HMI tags "Do_PLC"
   "System_okien_auto" : Bool = PLC HMI.System_okien_auto, 500 ms
   "Stopien_zasloniecia_rolet_manual" : Int = PLC HMI.Stopien_zasloniecia_rolet_manual, 100 ms
   "Przycisk_zraszania_manual" : Bool = PLC HMI.Przycisk_zraszacze_manual AT %Q0.2, 100 ms
   "Przycisk_wentylacja_manual" : Bool = PLC HMI.Przycisk_wentylacja_manual AT %Q0.1, 100 ms
   "Przycisk_grzanie_manual" : Bool = PLC HMI.Przycisk_grzanie_manual AT %Q0.0, 100 ms
   "Otwarcie_okien_man" : Bool = PLC HMI.Otwarcie_okien_manual AT %DB1.DBW0, 100 ms
   "Temperatura_auto" : Real = PLC HMI.Temperatura_auto, 500 ms
   "Naslonecznienie_auto" : Int = PLC HMI.Naslonecznienie_auto AT %DB1.DBW0, 500 ms
   "Wilgotnosc_powietrza_auto" : Int = PLC HMI.Wilgotnosc_powietrza_auto AT %DB1.DBW0, 500 ms
   "Wilgotnosc_gleby_auto" : Int = PLC HMI.Wilgotnosc_gleby_auto AT %DB1.DBW0, 500 ms
   "Przycisk_podlewania_manual" : Bool = PLC HMI.Przycisk_podlewanie_manual AT %Q0.2, 100 ms
   "Poziom_CO2_auto" : Int = PLC HMI.Poziom_CO2_auto AT %DB1.DBX0.0, 1 s

HMI tags "Z_PLC"
   "Czujnik_wilgotności_powietrza" : Int = PLC Wejscia_PLC.Czujnik_wilgotności_powietrza, 500 ms
   "Temperatura_wewnetrzna" : Real = PLC Wejscia_PLC.Temperatura_wewnetrzna, 500 ms
   "Czujnik_natezenia_światła" : Int = PLC Wejscia_PLC.Czujnik_natezenia_swiatła, 500 ms
   "Czujnik_wilgotności_gleby" : Int = PLC Wejscia_PLC.Czujnik_wilgotności_gleby, 500 ms
   "Wewnetrzny_czujnik_CO2" : Int = PLC Wejscia_PLC.Wewnetrzny_czujnik_CO2, 500 ms
   "Czujnik_wiatru" : Int = PLC Wejscia_PLC.Czujnik_wiatru, 500 ms
   "Stopien_zasloniecia_rolet" : Int = PLC Wejscia_PLC.Stopien_zasloniecia_rolet, 1 s
   "Zewnetrzny_czujnik_CO2" : Int = PLC Wejscia_PLC.Zewnetrzny_czujnik_CO2 AT %DB1.DBW0, 1 s
   "Temperatura_zewnetrzna" : Real = PLC Wejscia_PLC.Temperatura_zewnetrzna AT %DB1.DBW0, 1 s

discrete alarms
   6: 'Braku możliwości osiągnięcia wymaganego poziomu CO2 / Inability to reach required CO2 level / Unfähigkeit, erforderlichen CO2-Wert zu erreichen', class Warnings, trigger "Alarmy_alarm_word_DB" bit 0
   7: 'Zbyt niska temperatura utrzymuje się od dłuższego czasu. Sprawdź działanie grzałki / Temperature too low for extended period. Check heater operation. / Temperatur zu niedrig seit längerer Zeit. Heizung prüfen.', class Warnings, trigger "Alarmy_alarm_word_DB" bit 1
   8: 'Zbyt niska temperatura utrzymuje się od dłuższego czasu. Sprawdź działanie grzałki lub wentylatora / Temperature too low for extended period. Check heater or ventilator. / Temperatur zu niedrig seit längerer Zeit. Heizung oder Lüfter prüfen.', class Warnings, trigger "Alarmy_alarm_word_DB" bit 2

analog alarms
   1: 'Stężenie CO2 ma powyżej 1400 jednostek / CO2 concentration above 1400 units / CO2-Konzentration über 1400 Einheiten / Stężenie CO2 ma powyżej 1400 jednostek, dłużesze przebywanie w takim środowisku może być szkodliwe dla człowieka. Zalecane jest włączenie wentylacji lub otworzenie okien. / CO2 concentration above 1400 units, prolonged exposure may be harmful. Recommended to activate ventilation or open windows. / CO2-Konzentration über 1400 Einheiten, längere Exposition kann schädlich sein. Empfohlen: Lüftung aktivieren oder Fenster öffnen.', class Warnings, trigger "Wewnetrzny_czujnik_CO2"
   2: 'Temperatura powyżej 35 stopni / Temperature above 35 degrees / Temperatur über 35 Grad / Temperatura powyżej 35 stopni, zaleca się wyłączenie grzania. / Temperature above 35 degrees, recommended to turn off heating. / Temperatur über 35 Grad, empfohlen Heizung auszuschalten.', class Warnings, trigger "Temperatura_wewnetrzna"
   3: 'Podmuchy wiatru osiągają wartości powyżej 35 km/h, system automatyczny zamyka okna. / Wind gusts exceeding 35 km/h, automatic system closes windows. / Windböen über 35 km/h, automatisches System schließt Fenster.', class Warnings, trigger "Czujnik_wiatru"
   4: 'Stężenie CO2 ma powyżej 3000 jednostek. NIEZWŁOCZNIE OTWORZ OKNA ORAZ ZAŁĄCZ WENTYLATOR, NASTĘPNIE NALEŻY EWAKUOWAĆ WSZYSTKUCH ZNAJDUJĄCYCH SIĘ W POMIESZCZENIU / CO2 concentration above 3000 units. IMMEDIATELY OPEN WINDOWS AND TURN ON VENTILATOR, THEN EVACUATE ALL PERSONS FROM THE AREA. / CO2-Konzentration über 3000 Einheiten. SOFORT FENSTER ÖFFNEN UND LÜFTER EINSCHALTEN, DANN ALLE PERSONEN RÄUMEN. / Stężenie CO2 ma powyżej 3000 jednostek. NIEZWŁOCZNIE OTWORZ OKNA ORAZ ZAŁĄCZ WENTYLATOR, NASTĘPNIE NALEŻY EWAKUOWAĆ WSZYSTKUCH ZNAJDUJĄCYCH SIĘ W POMIESZCZENIU / CO2 concentration above 3000 units. IMMEDIATELY OPEN WINDOWS AND TURN ON VENTILATOR, THEN EVACUATE ALL PERSONS FROM THE AREA. / CO2-Konzentration über 3000 Einheiten. SOFORT FENSTER ÖFFNEN UND LÜFTER EINSCHALTEN, DANN ALLE PERSONEN RÄUMEN.', class Errors, trigger "Wewnetrzny_czujnik_CO2"
   5: 'Temperatura powyżej 45 stopni, NIEZWŁOCZNIE SPRAWDŹ DZIAŁANIE GRZAŁKI, TERMOMETRU LUB WENTYLATORA. / Temperature above 45 degrees, IMMEDIATELY CHECK HEATER, THERMOMETER OR VENTILATOR. / Temperatur über 45 Grad, SOFORT HEIZUNG, THERMOMETER ODER LÜFTER PRÜFEN. / Temperatura powyżej 45 stopni, NIEZWŁOCZNIE SPRAWDŹ DZIAŁANIE GRZAŁKI, TERMOMETRU LUB WENTYLATORA. JEŚLI TEMPERATURA NIE SPADA ZALECA SIĘ EWAKUOWAĆ WSZYSTKICH PRZEBYWAJĄCYCH W POMIESZCZENIU / Temperature above 45 degrees, IMMEDIATELY CHECK HEATER, THERMOMETER OR VENTILATOR. IF TEMPERATURE DOES NOT DROP, EVACUATE ALL PERSONS. / Temperatur über 45 Grad, SOFORT HEIZUNG, THERMOMETER ODER LÜFTER PRÜFEN. WENN TEMPERATUR NICHT SINKT, ALLE PERSONEN EVAKUIEREN.', class Errors, trigger "Temperatura_wewnetrzna"

recipe "Receptura_nr1": Temperatura <- "Tryb_auto_parametry_Temperatura", Wilgotność Powietrza <- "Tryb_auto_parametry_Wilgotnosc_powietrza", Wilgotność gleby <- "Tryb_auto_parametry_Wilgotnosc_gleby", System okien <- "Tryb_auto_parametry_System_okien", Stężenie CO2 <- "Tryb_auto_parametry_Stezenie_co2", Nasłonecznienie <- "Tryb_auto_parametry_Naslonecznienie"

screen "Root screen" 800x480, template "Template_1"
   on GenerateScreen: SetTag("Tag_ScreenNumber", 0)
   Button "Button_1" at 9,154 size 300x70; TextOff 'MANUAL MODE / TRYB MANUALNY / MANUELLER MODUS'
      on Click: ActivateScreen("tryb_manualny", 0)
   Button "Button_2" at 10,70 size 300x70; TextOff 'AUTOMATIC MODE / TRYB AUTOMATYCZNY / AUTOMATIKMODUS'
      on Click: ActivateScreen("tryb_automatyczny", 0)
   TextField "Text field_2" at 73,1 size 689x52; Text 'AUTOMATIC GREENHOUSE / AUTOMATYCZNA SZKLARNIA / AUTOMATISCHES GEWÄCHSHAUS'
   GraphicView "Graphic view_1" at 370,70 size 392x338; Picture "garden-tools-graphic-clipart-design-free-png"
   Button "Button_5" at 10,237 size 300x70; TextOff 'TRYB RECEPTUR / RECIPE MODE / REZEPTURMODUS'
      on Click: function_e3503463('\USB_X60.1\record.csv', U 0, 2, 1, N); ActivateScreen("Receptury", 0)
   Button "Button_3" at 10,322 size 300x70; TextOff 'SYMULACJA / SIMULATION'
      on Click: ActivateScreen("Symulacja_czujnikow", 0)

screen "tryb_manualny" 800x480
   on GenerateScreen: SetTag("Tag_ScreenNumber", 2)
   TextField "Text field_1" at 295,7 size 259x34; Text 'MANUAL MODE / TRYB MANUALNY / MANUELLER MODUS'
   TextField "Text field_4" at 511,174 size 171x23; Text 'WINDOW OPENING / OTWIERANIE OKIEN / FENSTERÖFFNUNG'
   Button "Button_4" at 518,261 size 80x70; TextOff 'WATERING / PODLEWANIE / BEWÄSSERUNG'
      on Click: InvertBit("Przycisk_podlewania_manual")
   Button "Button_5" at 611,261 size 80x70; TextOff 'HEATING / GRZANIE / HEIZUNG'
      on Click: InvertBit("Przycisk_grzanie_manual")
   Button "Button_6" at 701,261 size 80x70; TextOff 'VENTILATION / WENTYLACJA / LÜFTUNG'
      on Click: InvertBit("Przycisk_wentylacja_manual")
   GraphicView "Graphic view_1" at 710,356 size 60x60; Picture "fan_4829316"
      Visibility <- "Wentylator"
   GraphicView "Graphic view_6" at 622,356 size 60x60; Picture "heater_4463010"
      Visibility <- "Grzałka"
   GraphicView "Graphic view_7" at 527,356 size 64x60; Picture "irrigation_18631825"
      Visibility <- "Pompa_podlewanie"
   GraphicView "Graphic view_9" at 710,356 size 60x60; Picture "fan_off"
      Visibility <- "Wentylator"
   GraphicView "Graphic view_10" at 622,356 size 60x60; Picture "heater_off"
      Visibility <- "Grzałka"
   GraphicView "Graphic view_11" at 527,356 size 64x60; Picture "irrigation_off"
      Visibility <- "Pompa_podlewanie"
   Button "Button_14" at 6,7 size 43x43; TextOff 'HOME / DOM / HAUS'; PictureOff "home_1"
      on Click: ActivateScreen("Root screen", 0)
   Button "Button_1" at 740,0 size 60x60; TextOff 'Text'; PictureOff "Back_arrow"
      on Click: function_efd93a16()
   Circle "Circle_1" at 541,428 size 42x42
      Visibility <- "Pompa_podlewanie"
   Circle "Circle_4" at 541,428 size 42x42
      Visibility <- "Pompa_podlewanie"
   Circle "Circle_2" at 631,428 size 42x42
      Visibility <- "Grzałka"
   Circle "Circle_5" at 631,428 size 42x42
      Visibility <- "Grzałka"
   Circle "Circle_3" at 720,428 size 41x41
      Visibility <- "Wentylator"
   Circle "Circle_6" at 720,428 size 41x41
      Visibility <- "Wentylator"
   TextField "Text field_8" at 405,71 size 117x61; Text 'DEGREE OF BLINDS COVERAGE STOPIEŃ ZASŁONIECIA ROLET GRAD DER ROLLADEN- BEDECKUNG'
   Bar "Bar_6" at 624,82 size 165x66; MinimumValue 0; MaximumValue 100
      ProcessValue <- "Stopien_zasloniecia_rolet_manual"
   Button "Button_3" at 530,114 size 80x50; TextOff 'UNCOVER / ODSŁOŃ / ENTBLÖSSEN'
      on Click: function_b9b71300("Stopien_zasloniecia_rolet_manual", 5)
   Button "Button_7" at 530,60 size 80x50; TextOff 'COVER / ZASŁOŃ / ABDECKEN'
      on Press: function_dd21b452("Stopien_zasloniecia_rolet_manual", 5)
   Button "Button_2" at 425,261 size 80x70; TextOff 'MISTING / MIKROZRASZANIE / BESPRÜHUNG'
      on Click: InvertBit("Przycisk_zraszania_manual")
   GraphicView "Graphic view_2" at 434,356 size 60x60; Picture "sprinkler_4552152"
      Visibility <- "Pompa_zraszacze"
   GraphicView "Graphic view_3" at 434,356 size 60x60; Picture "sprinkler"
      Visibility <- "Pompa_zraszacze"
   Circle "Circle_7" at 443,428 size 42x42
      Visibility <- "Pompa_zraszacze"
   Circle "Circle_8" at 443,428 size 42x42
      Visibility <- "Pompa_zraszacze"
   Switch "Switch_1" at 499,199 size 209x37; CaptionText 'Schalter'; TextOff 'ZAMKNIĘTE / CLOSED / GESCHLOSSEN'; TextOn 'OTWARTE / OPEN / OFFEN'
      ProcessValue <- "Otwarcie_okien_man"
   TextField "Text field_3" at 11,375 size 212x23; Text 'WIND SPEED / SZYBKOŚĆ WIATRU / WINDGESCHWINDIGKEIT'
   IOField "I/O field_3" at 62,407 size 70x65; FormatPattern 999
      ProcessValue <- "Czujnik_wiatru"
   IOField "I/O field_1" at 48,189 size 101x32; FormatPattern 99999
      ProcessValue <- "Czujnik_natezenia_światła"
   TextField "Text field_15" at 129,408 size 52x72; Text 'Km h'
   IOField "I/O field_2" at 44,292 size 83x65; FormatPattern 9999
      ProcessValue <- "Wewnetrzny_czujnik_CO2"
   TextField "Text field_11" at 118,301 size 69x39; Text 'ppm'
   TextField "Text field_5" at 14,148 size 204x23; Text 'INSOLATION / NASŁONECZNIENIE / SONNENEINSTRAHLUNG'
   IOField "I/O field_8" at 58,95 size 93x40; FormatPattern 99.99
      ProcessValue <- "Temperatura_wewnetrzna"
   TextField "Text field_20" at 30,56 size 137x42; Text 'INTERIOR TEMPERATURE TEMPERATURA WEWNTĘTRZNA INNEN- TEMPERATUR'
   TextField "Text field_7" at 200,375 size 185x23; Text 'SOIL MOISTURE / WILGOTNOŚĆ GLEBY / BODENFEUCHTIGKEIT'
   IOField "I/O field_5" at 248,293 size 83x65; FormatPattern 9999
      ProcessValue <- "Zewnetrzny_czujnik_CO2"
   IOField "I/O field_4" at 266,174 size 69x65; FormatPattern 999
      ProcessValue <- "Czujnik_wilgotności_powietrza"
   IOField "I/O field_6" at 261,405 size 68x65; FormatPattern 999
      ProcessValue <- "Czujnik_wilgotności_gleby"
   TextField "Text field_12" at 324,182 size 47x46; Text '%'
   TextField "Text field_13" at 321,416 size 47x46; Text '%'
   TextField "Text field_16" at 325,302 size 69x39; Text 'ppm'
   IOField "I/O field_9" at 248,85 size 97x65; FormatPattern 99.99
      ProcessValue <- "Temperatura_zewnetrzna"
   TextField "Text field_23" at 333,90 size 46x46; Text '°C'
   TextField "Text field_22" at 229,57 size 132x42; Text 'EXTERIOR TEMPERATURE TEMPERATURA ZEWNĘTRZNA AUSSEN- TEMPERATUR'
   TextField "Text field_9" at 229,256 size 189x42; Text 'EXTERIOR CO2 CONCENTRATION ZEWNĘTRZNE STĘŻENIE CO2 AUSSEN- CO2-KONZENTRATION'
   TextField "Text field_6" at 180,143 size 128x42; Text 'AIR HUMIDITY WILGOTNOŚĆ POWIETRZA LUFT- FEUCHTIGKEIT'
   TextField "Text field_14" at 140,170 size 47x72; Text 'W m²'
   TextField "Text field_21" at 141,90 size 46x46; Text '°C'
   GraphicView "Graphic view_4" at 419,176 size 60x60; Picture "window_11250237"
   GraphicView "Graphic view_5" at 197,182 size 50x50; Picture "sensor_4212519"
   GraphicView "Graphic view_8" at 4,182 size 50x50; Picture "sensor_4212513"
   GraphicView "Graphic view_12" at 3,87 size 50x50; Picture "Thermometer_icon"
   GraphicView "Graphic view_13" at 199,87 size 50x50; Picture "Thermometer_icon"
   GraphicView "Graphic view_14" at 3,302 size 40x40; Picture "sensor_2828470"
   GraphicView "Graphic view_15" at 197,300 size 40x40; Picture "sensor_2828470"
   GraphicView "Graphic view_16" at 198,412 size 50x50; Picture "soil-sensor_11298794"
   GraphicView "Graphic view_17" at 3,416 size 50x50; Picture "anemometer_1113716"
   TextField "Text field_2" at 27,256 size 189x42; Text 'INTERIOR CO2 CONCENTRATION WEWNĘTRZNE STĘŻENIE CO2 INNEN- CO2-KONZENTRATION'

screen "praca" 800x480
   on GenerateScreen: SetTag("Tag_ScreenNumber", 5)
   GraphicView "Graphic view_4" at 275,402 size 70x70; Picture "soil-sensor_11298794"
   GraphicView "Graphic view_3" at 4,181 size 70x70; Picture "sensor_4212513"
   GraphicView "Graphic view_5" at 268,181 size 70x70; Picture "sensor_4212519"
   GraphicView "Graphic view_1" at 560,402 size 70x70; Picture "fan_4829316"
      Visibility <- "Wentylator"
   GraphicView "Graphic view_6" at 561,276 size 70x70; Picture "heater_4463010"
      Visibility <- "Grzałka"
   GraphicView "Graphic view_7" at 560,170 size 70x70; Picture "irrigation_18631825"
      Visibility <- "Pompa_podlewanie"
   GraphicView "Graphic view_8" at 12,403 size 70x70; Picture "anemometer_1113716"
   GraphicView "Graphic view_9" at 560,402 size 70x70; Picture "fan_off"
      Visibility <- "Wentylator"
   GraphicView "Graphic view_10" at 561,276 size 70x70; Picture "heater_off"
      Visibility <- "Grzałka"
   GraphicView "Graphic view_11" at 560,170 size 70x70; Picture "irrigation_off"
      Visibility <- "Pompa_podlewanie"
   GraphicView "Graphic view_12" at 279,273 size 70x70; Picture "sensor_2828470"
   TextField "Text field_1" at 53,158 size 204x23; Text 'INSOLATION / NASŁONECZNIENIE / SONNENEINSTRAHLUNG'
   TextField "Text field_3" at 45,379 size 212x23; Text 'WIND SPEED / SZYBKOŚĆ WIATRU / WINDGESCHWINDIGKEIT'
   TextField "Text field_5" at 290,158 size 223x23; Text 'AIR HUMIDITY / WILGOTNOŚĆ POWIETRZA / LUFTFEUCHTIGKEIT'
   TextField "Text field_6" at 319,379 size 185x23; Text 'SOIL MOISTURE / WILGOTNOŚĆ GLEBY / BODENFEUCHTIGKEIT'
   TextField "Text field_7" at 629,154 size 132x23; Text 'WATERING / PODLEWANIE / BEWÄSSERUNG'
   TextField "Text field_8" at 639,258 size 81x23; Text 'HEATING / GRZANIE / HEIZUNG'
   TextField "Text field_9" at 628,379 size 119x23; Text 'VENTILATION / WENTYLACJA / LÜFTUNG'
   TextField "Text field_10" at 80,10 size 256x34; Text 'LIVE PREVIEW / PODGLĄD NA ŻYWO / LIVE-VORSCHAU'
   Button "Button_1" at 750,0 size 50x50; TextOff 'BACK / WRÓĆ / ZURÜCK'; PictureOff "Back_arrow"
      on Click: function_efd93a16(); SetBit("HMI_Reset_Trybow")
   Button "Button_2" at 3,1 size 43x43; TextOff 'HOME / DOM / HAUS'; PictureOff "home_1"
      on Click: ActivateScreen("Root screen", 0); SetBit("HMI_Reset_Trybow")
   IOField "I/O field_3" at 95,408 size 70x65; FormatPattern 999
      ProcessValue <- "Czujnik_wiatru"
   IOField "I/O field_5" at 349,283 size 83x65; FormatPattern 9999
      ProcessValue <- "Zewnetrzny_czujnik_CO2"
   IOField "I/O field_4" at 378,178 size 69x65; FormatPattern 999
      ProcessValue <- "Czujnik_wilgotności_powietrza"
   IOField "I/O field_6" at 382,403 size 68x65; FormatPattern 999
      ProcessValue <- "Czujnik_wilgotności_gleby"
   TextField "Text field_12" at 447,196 size 47x46; Text '%'
   TextField "Text field_13" at 467,411 size 47x46; Text '%'
   TextField "Text field_14" at 193,170 size 47x72; Text 'W m²'
   IOField "I/O field_1" at 84,196 size 101x32; FormatPattern 99999
      ProcessValue <- "Czujnik_natezenia_światła"
   TextField "Text field_15" at 174,408 size 52x72; Text 'Km h'
   Circle "Circle_1" at 704,194 size 48x48
      Visibility <- "Pompa_podlewanie"
   Circle "Circle_2" at 703,289 size 48x48
      Visibility <- "Grzałka"
   TextField "Text field_16" at 448,289 size 69x39; Text 'ppm'
   Circle "Circle_4" at 704,194 size 48x48
      Visibility <- "Pompa_podlewanie"
   Circle "Circle_5" at 703,289 size 48x48
      Visibility <- "Grzałka"
   Circle "Circle_3" at 704,421 size 48x48
      Visibility <- "Wentylator"
   Circle "Circle_6" at 704,421 size 48x48
      Visibility <- "Wentylator"
   TextField "Text field_17" at 380,10 size 288x34; Text 'AUTOMATIC MODE / TRYB AUTOMATYCZNY / AUTOMATIKMODUS'
      Visibility <- "HMI_Aktywacja_trybu_automatycznego"
   GraphicView "Graphic view_13" at 561,69 size 70x70; Picture "sprinkler_4552152"
      Visibility <- "Pompa_zraszacze"
   GraphicView "Graphic view_14" at 561,69 size 70x70; Picture "sprinkler"
      Visibility <- "Pompa_zraszacze"
   Circle "Circle_7" at 704,89 size 48x48
      Visibility <- "Pompa_zraszacze"
   Circle "Circle_8" at 704,89 size 48x48
      Visibility <- "Pompa_zraszacze"
   TextField "Text field_19" at 613,58 size 156x23; Text 'MISTING / MIKROZRASZANIE / BESPRÜHUNG'
   GraphicView "Graphic view_15" at 1,72 size 70x70; Picture "Thermometer_icon"
   IOField "I/O field_8" at 74,79 size 97x65; FormatPattern 99.99
      ProcessValue <- "Temperatura_wewnetrzna"
   TextField "Text field_21" at 172,91 size 46x46; Text '°C'
   GraphicView "Graphic view_16" at 276,72 size 70x70; Picture "Thermometer_icon"
   IOField "I/O field_9" at 349,79 size 97x65; FormatPattern 99.99
      ProcessValue <- "Temperatura_zewnetrzna"
   TextField "Text field_23" at 448,88 size 46x46; Text '°C'
   TextField "Text field_20" at 59,55 size 137x42; Text 'INTERIOR TEMPERATURE TEMPERATURA WEWNTĘTRZNA INNEN- TEMPERATUR'
   TextField "Text field_22" at 336,55 size 132x42; Text 'EXTERIOR TEMPERATURE TEMPERATURA ZEWNĘTRZNA AUSSEN- TEMPERATUR'
   GraphicView "Graphic view_2" at 12,279 size 70x70; Picture "sensor_2828470"
   IOField "I/O field_2" at 82,289 size 83x65; FormatPattern 9999
      ProcessValue <- "Wewnetrzny_czujnik_CO2"
   TextField "Text field_11" at 181,295 size 69x39; Text 'ppm'
   TextField "Text field_2" at 84,258 size 189x42; Text 'INTERIOR CO2 CONCENTRATION WEWNĘTRZNE STĘŻENIE CO2 INNEN- CO2-KONZENTRATION'
   TextField "Text field_4" at 353,262 size 189x42; Text 'EXTERIOR CO2 CONCENTRATION ZEWNĘTRZNE STĘŻENIE CO2 AUSSEN- CO2-KONZENTRATION'
   TextField "Text field_18" at 381,10 size 230x34; Text 'TRYB RECEPTUR / RECIPE MODE / REZEPTURMODUS'
      Visibility <- "HMI_Aktywacja_trybu_Receptur"

Template "Template_1" 800x480
   Button "Exit" at 671,429 size 71x50; TextOn 'Exit / Beenden'; TextOff 'Exit / Beenden'; PictureOn "ExitRuntime_KTP700_Basic_PN_TR"; PictureOff "ExitRuntime_KTP700_Basic_PN_TR"
      on Release: StopRuntime(0)
   Button "Alarms" at 524,429 size 71x50; TextOn 'Alarms / Alarme'; TextOff 'Alarms / Alarme'; PictureOn "AlarmDisplay_KTP700_Basic_PN_TR"; PictureOff "AlarmDisplay_KTP700_Basic_PN_TR"
      on Release: function_ef3f5d25("Alarm window_Unacknowledged", -1)
   Button "Start screen" at 169,429 size 71x50; TextOn 'Start screen / Startbildschirm'; TextOff 'Start screen / Startbildschirm'; PictureOn "NavigateHome_KTP700_Basic_PN_TR"; PictureOff "NavigateHome_KTP700_Basic_PN_TR"
      on Release: ActivateScreen("Root screen", 0)
      Visibility <- "AlwaysTRUE"
   Button "Language" at 377,429 size 71x50; TextOn 'Language / Sprache'; TextOff 'Language / Sprache'; PictureOn "ToggleLanguage_KTP700_Basic_PN_TR"; PictureOff "ToggleLanguage_KTP700_Basic_PN_TR"
      on Release: function_fb9197e8(-1)

screen "Receptury" 800x480
   RecipeView "Recipe view_1" at 0,44 size 799x413; Recipe "Receptura_nr1"; RecipeNameCaption 'Select Recipe / Wybierz Recepturę / Rezept auswählen'; EntryNameCaption 'Saved Parameters / Zapisane Parametry / GespeParameter'; DataRecordNameCaption 'Select Recipe / Wybierz Recepturę / Rezept auswählen'
   GraphicView "Graphic view_1" at 529,157 size 35x35; Picture "Thermometer_icon"
   GraphicView "Graphic view_2" at 529,195 size 35x35; Picture "sensor_4212519"
   GraphicView "Graphic view_3" at 529,235 size 35x35; Picture "soil-sensor_11298794"
   GraphicView "Graphic view_4" at 529,274 size 35x35; Picture "window_11250237"
   GraphicView "Graphic view_5" at 529,313 size 35x35; Picture "sensor_2828470"
   GraphicView "Graphic view_6" at 529,353 size 35x35; Picture "sensor_4212513"
   TextField "Text field_11" at 569,155 size 39x38; Text '°C'
   TextField "Text field_18" at 569,195 size 39x38; Text '%'
   TextField "Text field_1" at 569,235 size 39x38; Text '%'
   TextField "Text field_2" at 564,274 size 48x32; Text '1/0'
   TextField "Text field_16" at 563,313 size 55x32; Text 'ppm'
   TextField "Text field_6" at 576,344 size 25x50; Text 'W m'
   TextField "Text field_3" at 593,367 size 22x17; Text '2 / 2.0'
   Button "Button_1" at 750,0 size 50x50; TextOff 'BACK / WRÓĆ / ZURÜCK'; PictureOff "Back_arrow"
      on Click: function_efd93a16()
   Button "Button_14" at 3,1 size 43x43; TextOff 'HOME / DOM / HAUS'; PictureOff "home_1"
      on Click: ActivateScreen("Root screen", 0)
   TextField "Text field_4" at 320,2 size 189x37; Text 'RECEPTURY / RECIPES / REZEPTUREN'
   TextField "Text field_5" at 12,448 size 50x23; Text 'Nowy / New / Neu'
   TextField "Text field_7" at 69,448 size 85x23; Text 'Zapisz / Save / Speichern'
   TextField "Text field_8" at 137,448 size 70x23; Text 'Usuń / Delete / Löschen'
   TextField "Text field_9" at 197,444 size 53x36; Text 'Zmień Nazwę Change Name Ändere Namen'
   TextField "Text field_10" at 672,444 size 62x36; Text 'Załaduj z PLC Load from PLC Lade von PLC'
   TextField "Text field_12" at 735,444 size 52x36; Text 'Załaduj do PLC Load to PLC Lade in PLC'
   Button "Button_2" at 379,406 size 281x40; TextOff 'ZATWIERDŹ / CONFIRM / BESTÄTIGEN'
      on Click: ResetBit("HMI_Reset_Trybow"); SetBit("HMI_Aktywacja_trybu_Receptur"); ActivateScreen("praca", 0)
   TextField "Text field_13" at 435,450 size 246x23; Text 'Przejdź w tryb pracy / Switch to operation mode / Zum Betriebsmodus wechseln'
   Button "Button_3" at 282,407 size 50x40; TextOff 'Z / From / Von'; PictureOff "Graphic_9"
      on Click: function_ea909784(1, U 0, '\USB_X60.1\record.csv', 2, 1, N)
   TextField "Text field_14" at 263,444 size 109x36; Text 'Zapisz Kopię zapasową Save Backup Copy Sichere Backup- Kopie'

screen "Symulacja_czujnikow" 800x480
   TextField "Text field_1" at 12,58 size 252x23; Text 'Czujnik Wilgotności powietrza / Air humidity sensor / Luftfeuchtigkeitssensor'
   TextField "Text field_2" at 306,58 size 215x23; Text 'Czujnik Wilgotności gleby / Soil moisture sensor / Bodenfeuchtigkeitssensor'
   TextField "Text field_3" at 32,202 size 202x23; Text 'Termometr wewnętrzny / Internal thermometer / Innenthermometer'
   TextField "Text field_4" at 323,202 size 197x23; Text 'Termometr zewnętrzny / External thermometer / Außenthermometer'
   TextField "Text field_5" at 566,58 size 216x23; Text 'Czujnik natężenia światła / Light intensity sensor / Lichtintensitätssensor'
   TextField "Text field_6" at 607,202 size 124x23; Text 'Czujnik wiatru / Wind sensor / Windsensor'
   TextField "Text field_7" at 27,346 size 208x23; Text 'Wewnętrzny czujnik CO2 / Internal CO2 sensor / Interner CO2-Sensor'
   TextField "Text field_8" at 306,346 size 202x23; Text 'Zewnętrzny czujnik CO2 / External CO2 sensor / Externer CO2-Sensor'
   TextField "Text field_9" at 569,346 size 210x23; Text 'Stopień zasłonięcia rolet / Degree of blind coverage / Rolladenabdeckungsgrad'
   IOField "I/O field_4" at 599,94 size 150x60; FormatPattern 9999
      ProcessValue <- "Czujnik_natezenia_światła"
   IOField "I/O field_5" at 599,242 size 150x60; FormatPattern 999
      ProcessValue <- "Czujnik_wiatru"
   IOField "I/O field_6" at 69,375 size 150x60; FormatPattern 9999
      ProcessValue <- "Wewnetrzny_czujnik_CO2"
   IOField "I/O field_7" at 346,375 size 150x60; FormatPattern 9999
      ProcessValue <- "Zewnetrzny_czujnik_CO2"
   IOField "I/O field_8" at 599,375 size 150x60; FormatPattern 999
      ProcessValue <- "Stopien_zasloniecia_rolet"
   IOField "I/O field_10" at 69,94 size 150x60; FormatPattern 999
      ProcessValue <- "Czujnik_wilgotności_powietrza"
   IOField "I/O field_11" at 346,94 size 150x60; FormatPattern 999
      ProcessValue <- "Czujnik_wilgotności_gleby"
   IOField "I/O field_12" at 69,242 size 150x60; FormatPattern 99.9
      ProcessValue <- "Temperatura_wewnetrzna"
   IOField "I/O field_13" at 346,242 size 150x60; FormatPattern 99.9
      ProcessValue <- "Temperatura_zewnetrzna"
   TextField "Text field_10" at 248,5 size 321x34; Text 'SENSOR SIMULATION / SYMULACJA CZUJNIKÓW / SENSOR-SIMULATION'
   Button "Button_1" at 750,0 size 50x50; TextOff 'BACK / WRÓĆ / ZURÜCK'; PictureOff "Back_arrow"
      on Click: function_efd93a16()
   Button "Button_14" at 3,1 size 43x43; TextOff 'HOME / DOM / HAUS'; PictureOff "home_1"
      on Click: ActivateScreen("Root screen", 0)

screen "tryb_automatyczny" 800x480
   on GenerateScreen: SetTag("Tag_ScreenNumber", 1)
   IOField "I/O field_1" at 67,322 size 57x40; FormatPattern 99.9
      ProcessValue <- "Temperatura_wewnetrzna"
   Button "Button_1" at 745,0 size 55x55; TextOff 'BACK / WRÓĆ / ZURÜCK'; PictureOff "Back_arrow"
      on Click: function_efd93a16()
   Button "Button_2" at 373,382 size 416x89; TextOff 'CONFIRM / ZATWIERDŹ / BESTÄTIGEN'
      on Click: ResetBit("HMI_Reset_Trybow"); SetBit("HMI_Aktywacja_trybu_automatycznego"); ActivateScreen("praca", 0)
   Bar "Bar_1" at 7,110 size 50x250; MinimumValue 0; MaximumValue 45
      ProcessValue <- "Temperatura_auto"
   TextField "Text field_2" at 1,71 size 132x23; Text 'TEMPERATURE / TEMPERATURA / TEMPERATUR'
   Bar "Bar_2" at 170,111 size 50x250; MinimumValue 0; MaximumValue 100
      ProcessValue <- "Wilgotnosc_powietrza_auto"
   TextField "Text field_3" at 165,68 size 138x42; Text 'AIR HUMIDITY WILGOTNOŚĆ POWIETRZA LUFT- FEUCHTIGKEIT'
   Button "Button_3" at 71,115 size 75x45; TextOff '+0.5 °C'
      on Press: function_dd21b452("Temperatura_auto", 0.5)
   Button "Button_7" at 71,183 size 75x45; TextOff '-0.5 °C'
      on Press: function_b9b71300("Temperatura_auto", 0.5)
   IOField "I/O field_2" at 67,251 size 62x40; FormatPattern 99.9
      ProcessValue <- "Temperatura_auto"
   TextField "Text field_11" at 122,260 size 23x22; Text '°C'
   TextField "Text field_9" at 122,333 size 23x22; Text '°C'
   Bar "Bar_4" at 335,111 size 50x250; MinimumValue 0; MaximumValue 100
      ProcessValue <- "Wilgotnosc_gleby_auto"
   TextField "Text field_10" at 332,65 size 158x42; Text 'SOIL MOISTURE WILGOTNOŚĆ GLEBY BODEN- FEUCHTIGKEIT'
   Button "Button_8" at 398,132 size 65x40; TextOff '+2%'
      on Click: function_dd21b452("Wilgotnosc_gleby_auto", 2)
   Button "Button_9" at 398,181 size 65x40; TextOff '-0.02 / -2%'
      on Click: function_b9b71300("Wilgotnosc_gleby_auto", 2)
   IOField "I/O field_5" at 402,255 size 60x40; FormatPattern 999
      ProcessValue <- "Wilgotnosc_gleby_auto"
   IOField "I/O field_6" at 404,325 size 58x40; FormatPattern 999
      ProcessValue <- "Czujnik_wilgotności_gleby"
   TextField "Text field_12" at 385,243 size 108x22; Text 'SET / USTAWIONA / EINGESTELLT'
   TextField "Text field_13" at 389,314 size 86x22; Text 'ACTUAL / AKTUALNA / AKTUELL'
   TextField "Text field_14" at 439,264 size 23x22; Text '%'
   TextField "Text field_15" at 439,335 size 23x22; Text '%'
   Button "Button_10" at 229,126 size 65x40; TextOff '+5%'
      on Click: function_dd21b452("Wilgotnosc_powietrza_auto", 5)
   Button "Button_11" at 229,186 size 65x40; TextOff '-0.05 / -5%'
      on Click: function_b9b71300("Wilgotnosc_powietrza_auto", 5)
   IOField "I/O field_4" at 234,254 size 66x40; FormatPattern 999
      ProcessValue <- "Wilgotnosc_powietrza_auto"
   IOField "I/O field_7" at 236,320 size 62x40; FormatPattern 999
      ProcessValue <- "Czujnik_wilgotności_powietrza"
   TextField "Text field_16" at 223,241 size 108x22; Text 'SET / USTAWIONA / EINGESTELLT'
   TextField "Text field_17" at 223,306 size 86x22; Text 'ACTUAL / AKTUALNA / AKTUELL'
   TextField "Text field_18" at 275,263 size 23x22; Text '%'
   TextField "Text field_19" at 275,328 size 23x22; Text '%'
   Button "Button_14" at 4,7 size 45x45; TextOff 'HOME / DOM / HAUS'; PictureOff "home_1"
      on Click: ActivateScreen("Root screen", 0)
   TextField "Text field_4" at 143,381 size 151x23; Text 'WINDOW SYSTEM / SYSTEM OKIEN / FENSTERSYSTEM'
   Switch "Switch_1" at 106,410 size 216x46; TextOn 'EIN'; CaptionText 'Schalter'; TextOff 'AUS'
      ProcessValue <- "System_okien_auto"
   GraphicView "Graphic view_1" at 129,70 size 40x40; Picture "Thermometer_icon"
   GraphicView "Graphic view_2" at 281,68 size 40x40; Picture "sensor_4212519"
   TextField "Text field_5" at 60,309 size 86x22; Text 'ACTUAL / AKTUALNA / AKTUELL'
   TextField "Text field_6" at 57,237 size 108x22; Text 'SET / USTAWIONA / EINGESTELLT'
   GraphicView "Graphic view_3" at 443,71 size 40x40; Picture "soil-sensor_11298794"
   TextField "Text field_1" at 255,4 size 291x47; Text 'TRYB AUTOMATYCZNY / AUTOMATIC MODE / AUTOMATIKMODUS'
   Bar "Bar_3" at 496,111 size 50x250; MinimumValue 0; MaximumValue 1500
      ProcessValue <- "Naslonecznienie_auto"
   TextField "Text field_7" at 488,55 size 194x22; Text 'INSOLATION / NASŁONECZNIENIE / SONNENEINSTRAHLUNG'
   GraphicView "Graphic view_4" at 585,86 size 40x40; Picture "sensor_4212513"
   Button "Button_4" at 553,131 size 82x43; TextOff '+50 W m'
      on Click: function_dd21b452("Naslonecznienie_auto", 50)
   Button "Button_5" at 554,186 size 82x43; TextOff '-50 W m'
      on Click: function_b9b71300("Naslonecznienie_auto", 50)
   IOField "I/O field_3" at 561,254 size 61x40; FormatPattern 9999
      ProcessValue <- "Naslonecznienie_auto"
   TextField "Text field_8" at 545,242 size 108x22; Text 'SET / USTAWIONE / EINGESTELLT'
   IOField "I/O field_8" at 563,325 size 62x40; FormatPattern 9999
      ProcessValue <- "Czujnik_natezenia_światła"
   TextField "Text field_20" at 549,313 size 85x22; Text 'ACTUAL / AKTUALNE / AKTUELLE'
   TextField "Text field_23" at 616,150 size 25x18; Text '2 / 2.0'
   TextField "Text field_24" at 614,205 size 25x18; Text '2 / 2.0'
   Bar "Bar_5" at 652,110 size 45x250; MinimumValue 400; MaximumValue 950
      ProcessValue <- "Poziom_CO2_auto"
   TextField "Text field_21" at 656,65 size 109x23; Text 'CO2 LEVEL / POZIOM CO2 / CO2-PEGEL'
   IOField "I/O field_9" at 723,254 size 66x40; FormatPattern 999
      ProcessValue <- "Poziom_CO2_auto"
   TextField "Text field_22" at 692,241 size 108x22; Text 'SET / USTAWIONY / EINGESTELLT'
   IOField "I/O field_10" at 723,333 size 62x40; FormatPattern 999
      ProcessValue <- "Wewnetrzny_czujnik_CO2"
   TextField "Text field_25" at 708,314 size 86x22; Text 'ACTUAL / AKTUALNA / AKTUELL'
   Button "Button_6" at 714,134 size 73x40; TextOff '+25ppm'
      on Click: function_dd21b452("Poziom_CO2_auto", 25)
   Button "Button_12" at 714,186 size 73x40; TextOff '-25ppm'
      on Click: function_b9b71300("Poziom_CO2_auto", 25)
   GraphicView "Graphic view_5" at 754,83 size 40x40; Picture "sensor_2828470"
   GraphicView "Graphic view_6" at 17,400 size 55x55; Picture "window_11250237"
*)